(* Logix 5000 project; controller NWGG 1756-L72 rev 35.12; software revision 35.00; part 11 of 19 *)
(* tags used below, declared in another part *)
   _108M : ALIAS FOR O25[10].15;
   _109M : ALIAS FOR O25[10].9;
   _116M : ALIAS FOR O25[10].10;
   _117M : ALIAS FOR O25[10].8;
   _11_GATE_PO1 : ALIAS FOR N14[11];
   _11_GATE_PO_STOR : REAL;
   _123M : ALIAS FOR O25[10].6;
   _12_GATE_PO1 : ALIAS FOR N14[12];
   _12_GATE_PO_STOR : REAL;
   _13_GATE_PO1 : ALIAS FOR N14[13];
   _13_GATE_PO_STOR : REAL;
   _14_GATE_PO1 : ALIAS FOR N14[14];
   _14_GATE_PO_STOR : REAL;
   _15_GATE_PO1 : ALIAS FOR N14[15];
   _15_GATE_PO_STOR : REAL;
   _16_GATE_PO1 : ALIAS FOR N14[16];
   _16_GATE_PO_STOR : REAL;
   _17_GATE_PO1 : ALIAS FOR N14[17];
   _17_GATE_PO_STOR : REAL;
   _21_GATE_PO1 : ALIAS FOR N14[21];
   _21_GATE_PO_STOR : REAL;
   _22_GATE_PO1 : ALIAS FOR N14[22];
   _22_GATE_PO_STOR : REAL;
   _23_GATE_PO1 : ALIAS FOR N14[23];
   _23_GATE_PO_STOR : REAL;
   _24_GATE_PO1 : ALIAS FOR N14[24];
   _24_GATE_PO_STOR : REAL;
   _25_GATE_PO1 : ALIAS FOR N14[25];
   _25_GATE_PO_STOR : REAL;
   _26_GATE_PO1 : ALIAS FOR N14[26];
   _26_GATE_PO_STOR : REAL;
   _35M : ALIAS FOR O25[10].13;
   _43M : ALIAS FOR O25[10].14;
   _705M : ALIAS FOR O25[10].12;
   B3 : DINT[250];
   cpBinGateRates : DINT[50];
   cpBINOPEN : DINT;
   cpCleanBulk : BOOL;
   cpTicketBinActive : DINT;
   cpTicketBinSet : DINT;
   cpVAR_BINARRAY : STRING[50];
   cpVAR_CNT_ONS : DINT;
   cpVarTrimTemp : STRING;
   indexTbl : DINT;
   indexTRTTbl : DINT;
   O24 : INT[32];
   O24_007_Bit10 : ALIAS FOR O24[7].10;
   O24_007_Bit11 : ALIAS FOR O24[7].11;
   O24_007_Bit12 : ALIAS FOR O24[7].12;
   O24_007_Bit13 : ALIAS FOR O24[7].13;
   O24_007_Bit14 : ALIAS FOR O24[7].14;
   P10_RUN_AU1 : ALIAS FOR B3[4].10;
   P1_RUN_AUT1 : ALIAS FOR B3[4].1;
   P2_RUN_AUT1 : ALIAS FOR B3[4].2;
   P3_RUN_AUT1 : ALIAS FOR B3[4].3;
   P4_RUN_AUT1 : ALIAS FOR B3[4].4;
   P5_RUN_AUT1 : ALIAS FOR B3[4].5;
   P6_RUN_AUT1 : ALIAS FOR B3[4].6;
   P7_RUN_AUT1 : ALIAS FOR B3[4].7;
   P8_RUN_AUT1 : ALIAS FOR B3[4].8;
   PUMP_13_RUN : ALIAS FOR R3M1_AENTR:3:O.8;
   PUMP_14_RUN : ALIAS FOR R3M1_AENTR:3:O.9;
   PUMP_15_RUN : ALIAS FOR R3M1_AENTR:3:O.14;
   spBinGateRates : DINT[50];
   spTicketProcessing : BOOL;
   strEmptyVar : STRING;
   TicketTreatPumpActive : DINT;
   TicketTreatPumpSet : DINT;
   TRT_ARRAY : STRING[50];
   TRT_CNT : DINT;
   TRT_CNT_ONS : DINT;
   Trt_CntStore : DINT;
   TRT_PumpRATE : DINT[50];
   TRT_TICKETtable : STRING[100];
   TRT_TickettableItemNo : DINT[50];
   TRT_TICKETtableRate : DINT[100];
   TrtTrimTemp : STRING;
   VAR_CNT : DINT;
   Var_CntStore : DINT;
   VAR_TICKETtable : STRING[20];
   VAR_TickettableItemNo : DINT[50];
   VAR_TICKETtableRate : DINT[100];
   vartableONS : DINT;
   zzztmpTANKtest : DINT[10];
(* MainProgram, continued *)

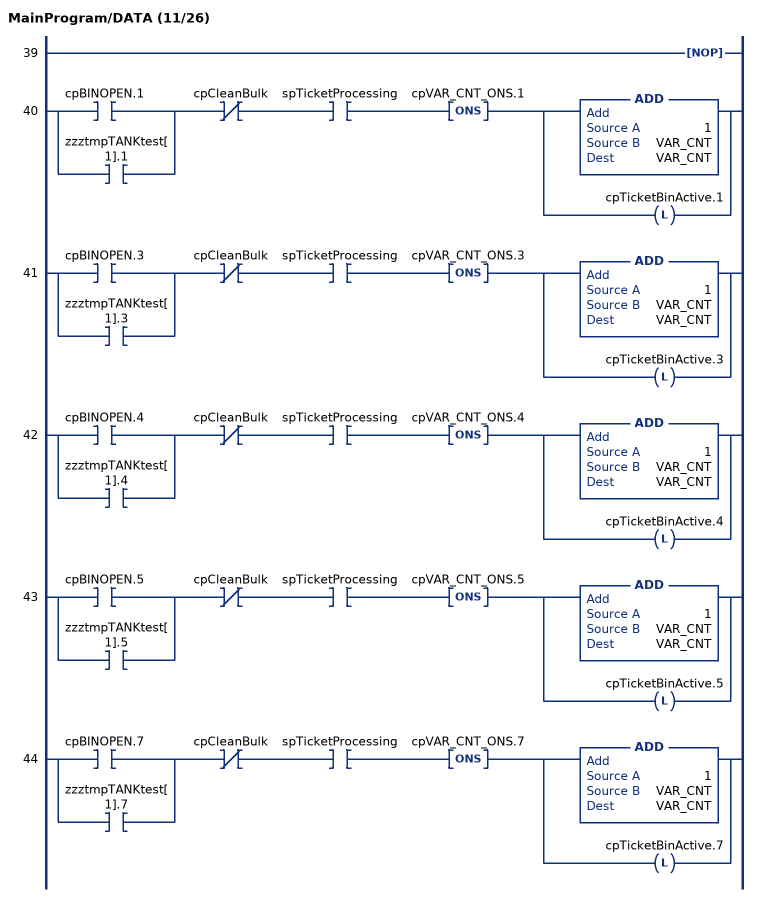
   [picture p209: MainProgram/DATA rungs 39-44]
   39: NOP();
   40: [XIC(cpBINOPEN.1) ,XIC(zzztmpTANKtest[1].1) ]XIO(cpCleanBulk)XIC(spTicketProcessing)ONS(cpVAR_CNT_ONS.1)[ADD(1,VAR_CNT,VAR_CNT) ,OTL(cpTicketBinActive.1) ];
   41: [XIC(cpBINOPEN.3) ,XIC(zzztmpTANKtest[1].3) ]XIO(cpCleanBulk)XIC(spTicketProcessing)ONS(cpVAR_CNT_ONS.3)[ADD(1,VAR_CNT,VAR_CNT) ,OTL(cpTicketBinActive.3) ];
   42: [XIC(cpBINOPEN.4) ,XIC(zzztmpTANKtest[1].4) ]XIO(cpCleanBulk)XIC(spTicketProcessing)ONS(cpVAR_CNT_ONS.4)[ADD(1,VAR_CNT,VAR_CNT) ,OTL(cpTicketBinActive.4) ];
   43: [XIC(cpBINOPEN.5) ,XIC(zzztmpTANKtest[1].5) ]XIO(cpCleanBulk)XIC(spTicketProcessing)ONS(cpVAR_CNT_ONS.5)[ADD(1,VAR_CNT,VAR_CNT) ,OTL(cpTicketBinActive.5) ];
   44: [XIC(cpBINOPEN.7) ,XIC(zzztmpTANKtest[1].7) ]XIO(cpCleanBulk)XIC(spTicketProcessing)ONS(cpVAR_CNT_ONS.7)[ADD(1,VAR_CNT,VAR_CNT) ,OTL(cpTicketBinActive.7) ];
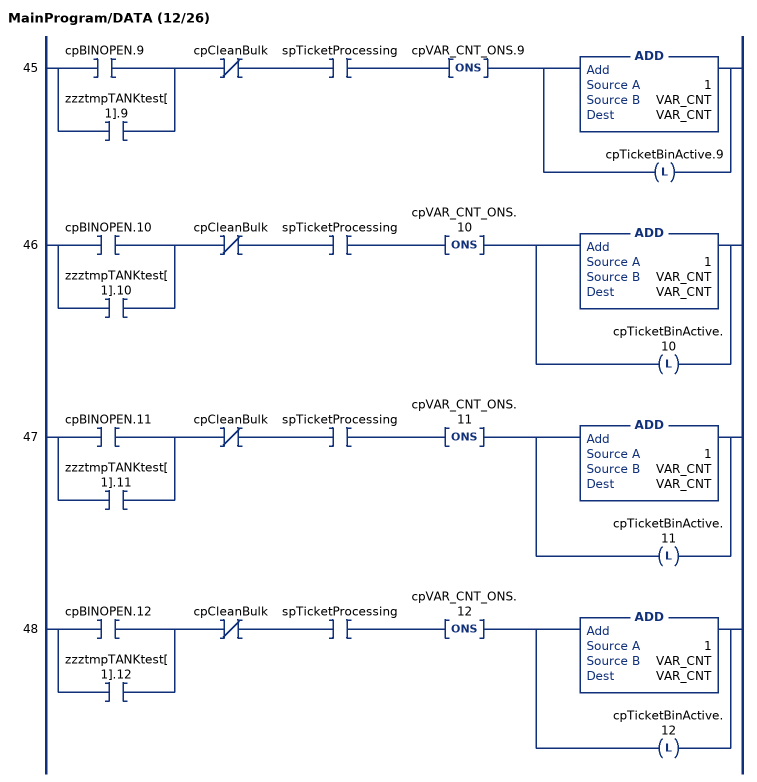
   45: [XIC(cpBINOPEN.9) ,XIC(zzztmpTANKtest[1].9) ]XIO(cpCleanBulk)XIC(spTicketProcessing)ONS(cpVAR_CNT_ONS.9)[ADD(1,VAR_CNT,VAR_CNT) ,OTL(cpTicketBinActive.9) ];
   46: [XIC(cpBINOPEN.10) ,XIC(zzztmpTANKtest[1].10) ]XIO(cpCleanBulk)XIC(spTicketProcessing)ONS(cpVAR_CNT_ONS.10)[ADD(1,VAR_CNT,VAR_CNT) ,OTL(cpTicketBinActive.10) ];
   47: [XIC(cpBINOPEN.11) ,XIC(zzztmpTANKtest[1].11) ]XIO(cpCleanBulk)XIC(spTicketProcessing)ONS(cpVAR_CNT_ONS.11)[ADD(1,VAR_CNT,VAR_CNT) ,OTL(cpTicketBinActive.11) ];
   48: [XIC(cpBINOPEN.12) ,XIC(zzztmpTANKtest[1].12) ]XIO(cpCleanBulk)XIC(spTicketProcessing)ONS(cpVAR_CNT_ONS.12)[ADD(1,VAR_CNT,VAR_CNT) ,OTL(cpTicketBinActive.12) ];
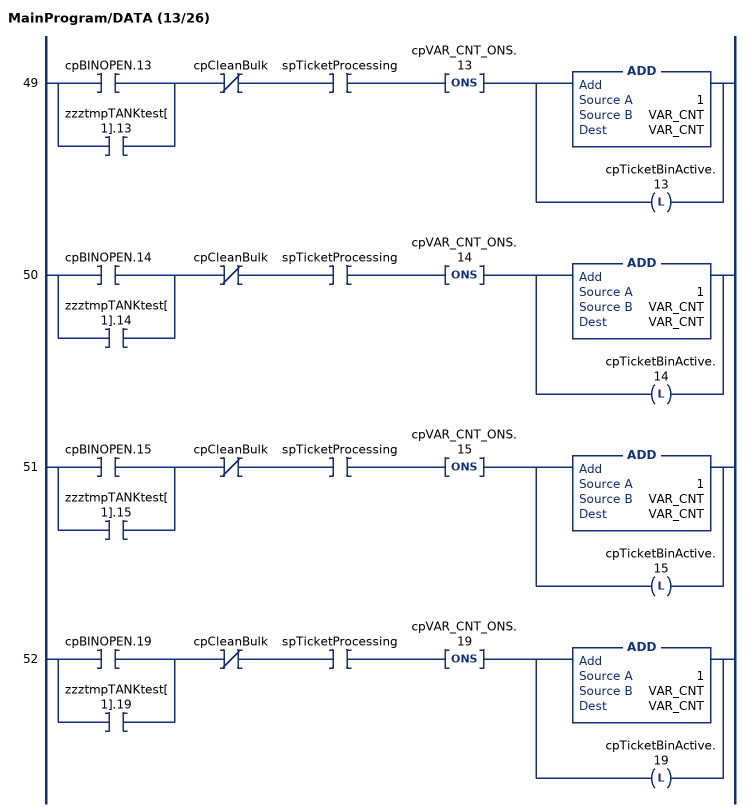
   49: [XIC(cpBINOPEN.13) ,XIC(zzztmpTANKtest[1].13) ]XIO(cpCleanBulk)XIC(spTicketProcessing)ONS(cpVAR_CNT_ONS.13)[ADD(1,VAR_CNT,VAR_CNT) ,OTL(cpTicketBinActive.13) ];
   50: [XIC(cpBINOPEN.14) ,XIC(zzztmpTANKtest[1].14) ]XIO(cpCleanBulk)XIC(spTicketProcessing)ONS(cpVAR_CNT_ONS.14)[ADD(1,VAR_CNT,VAR_CNT) ,OTL(cpTicketBinActive.14) ];
   51: [XIC(cpBINOPEN.15) ,XIC(zzztmpTANKtest[1].15) ]XIO(cpCleanBulk)XIC(spTicketProcessing)ONS(cpVAR_CNT_ONS.15)[ADD(1,VAR_CNT,VAR_CNT) ,OTL(cpTicketBinActive.15) ];
   52: [XIC(cpBINOPEN.19) ,XIC(zzztmpTANKtest[1].19) ]XIO(cpCleanBulk)XIC(spTicketProcessing)ONS(cpVAR_CNT_ONS.19)[ADD(1,VAR_CNT,VAR_CNT) ,OTL(cpTicketBinActive.19) ];
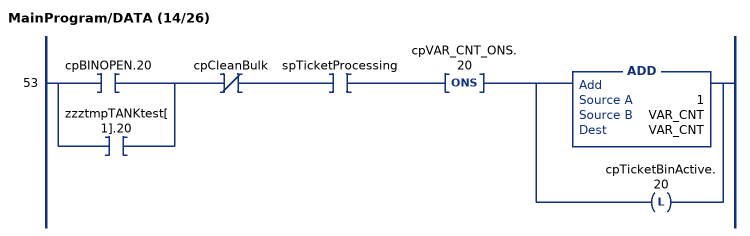
   53: [XIC(cpBINOPEN.20) ,XIC(zzztmpTANKtest[1].20) ]XIO(cpCleanBulk)XIC(spTicketProcessing)ONS(cpVAR_CNT_ONS.20)[ADD(1,VAR_CNT,VAR_CNT) ,OTL(cpTicketBinActive.20) ];
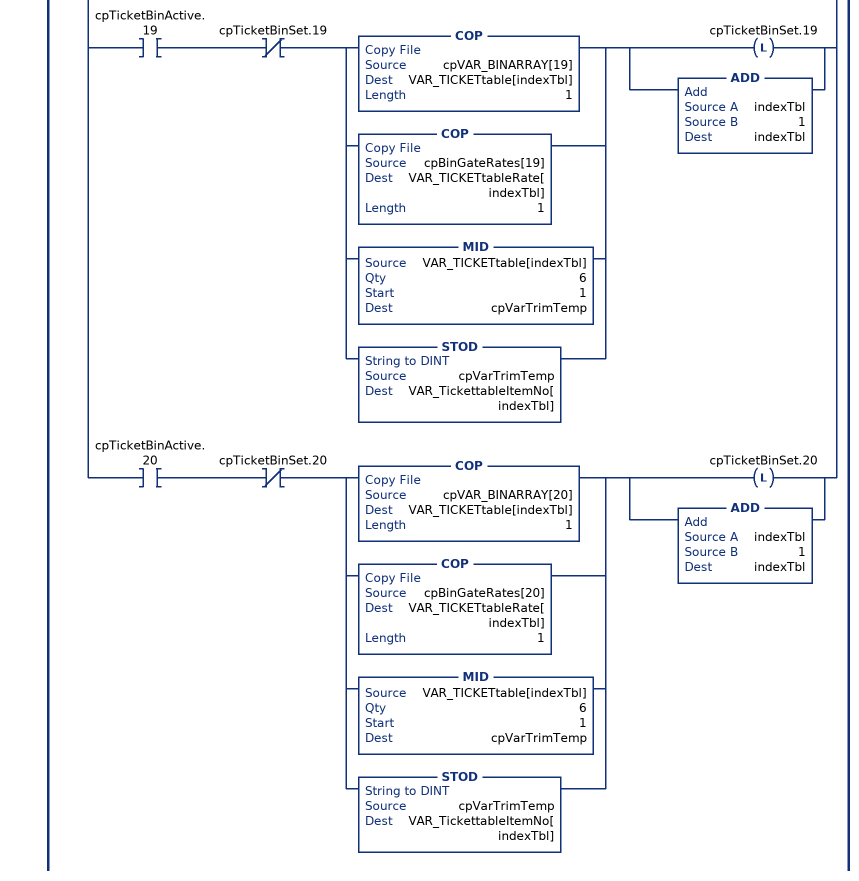
   54: GRT(VAR_CNT,0)LES(indexTbl,VAR_CNT)[XIC(cpTicketBinActive.1) XIO(cpTicketBinSet.1) [COP(cpVAR_BINARRAY[1],VAR_TICKETtable[indexTbl],1) ,COP(cpBinGateRates[1],VAR_TICKETtableRate[indexTbl],1) ,MID(VAR_TICKETtable[indexTbl],6,1,cpVarTrimTemp) ,STOD(cpVarTrimTemp,VAR_TickettableItemNo[indexTbl]) ] [OTL(cpTicketBinSet.1) ,ADD(indexTbl,1,indexTbl) ] ,XIC(cpTicketBinActive.3) XIO(cpTicketBinSet.3) [COP(cpVAR_BINARRAY[3],VAR_TICKETtable[indexTbl],1) ,COP(cpBinGateRates[3],VAR_TICKETtableRate[indexTbl],1) ,MID(VAR_TICKETtable[indexTbl],6,1,cpVarTrimTemp) ,STOD(cpVarTrimTemp,VAR_TickettableItemNo[indexTbl]) ] [OTL(cpTicketBinSet.3) ,ADD(indexTbl,1,indexTbl) ] ,XIC(cpTicketBinActive.4) XIO(cpTicketBinSet.4) [COP(cpVAR_BINARRAY[4],VAR_TICKETtable[indexTbl],1) ,COP(cpBinGateRates[4],VAR_TICKETtableRate[indexTbl],1) ,MID(VAR_TICKETtable[indexTbl],6,1,cpVarTrimTemp) ,STOD(cpVarTrimTemp,VAR_TickettableItemNo[indexTbl]) ] [OTL(cpTicketBinSet.4) ,ADD(indexTbl,1,indexTbl) ] ,XIC(cpTicketBinActive.5) XIO(cpTicketBinSet.5) [COP(cpVAR_BINARRAY[5],VAR_TICKETtable[indexTbl],1) ,COP(cpBinGateRates[5],VAR_TICKETtableRate[indexTbl],1) ,MID(VAR_TICKETtable[indexTbl],6,1,cpVarTrimTemp) ,STOD(cpVarTrimTemp,VAR_TickettableItemNo[indexTbl]) ] [OTL(cpTicketBinSet.5) ,ADD(indexTbl,1,indexTbl) ] ,XIC(cpTicketBinActive.7) XIO(cpTicketBinSet.7) [COP(cpVAR_BINARRAY[7],VAR_TICKETtable[indexTbl],1) ,COP(cpBinGateRates[7],VAR_TICKETtableRate[indexTbl],1) ,MID(VAR_TICKETtable[indexTbl],6,1,cpVarTrimTemp) ,STOD(cpVarTrimTemp,VAR_TickettableItemNo[indexTbl]) ] [OTL(cpTicketBinSet.7) ,ADD(indexTbl,1,indexTbl) ] ,XIC(cpTicketBinActive.9) XIO(cpTicketBinSet.9) [COP(cpVAR_BINARRAY[9],VAR_TICKETtable[indexTbl],1) ,COP(cpBinGateRates[9],VAR_TICKETtableRate[indexTbl],1) ,MID(VAR_TICKETtable[indexTbl],6,1,cpVarTrimTemp) ,STOD(cpVarTrimTemp,VAR_TickettableItemNo[indexTbl]) ] [OTL(cpTicketBinSet.9) ,ADD(indexTbl,1,indexTbl) ] ,XIC(cpTicketBinActive.10) XIO(cpTicketBinSet.10) [COP(cpVAR_BINARRAY[10],VAR_TICKETtable[indexTbl],1) ,COP(cpBinGateRates[10],VAR_TICKETtableRate[indexTbl],1) ,MID(VAR_TICKETtable[indexTbl],6,1,cpVarTrimTemp) ,STOD(cpVarTrimTemp,VAR_TickettableItemNo[indexTbl]) ] [OTL(cpTicketBinSet.10) ,ADD(indexTbl,1,indexTbl) ] ,XIC(cpTicketBinActive.11) XIO(cpTicketBinSet.11) [COP(cpVAR_BINARRAY[11],VAR_TICKETtable[indexTbl],1) ,COP(cpBinGateRates[11],VAR_TICKETtableRate[indexTbl],1) ,MID(VAR_TICKETtable[indexTbl],6,1,cpVarTrimTemp) ,STOD(cpVarTrimTemp,VAR_TickettableItemNo[indexTbl]) ] [OTL(cpTicketBinSet.11) ,ADD(indexTbl,1,indexTbl) ] ,XIC(cpTicketBinActive.12) XIO(cpTicketBinSet.12) [COP(cpVAR_BINARRAY[12],VAR_TICKETtable[indexTbl],1) ,COP(cpBinGateRates[12],VAR_TICKETtableRate[indexTbl],1) ,MID(VAR_TICKETtable[indexTbl],6,1,cpVarTrimTemp) ,STOD(cpVarTrimTemp,VAR_TickettableItemNo[indexTbl]) ] [OTL(cpTicketBinSet.12) ,ADD(indexTbl,1,indexTbl) ] ,XIC(cpTicketBinActive.13) XIO(cpTicketBinSet.13) [COP(cpVAR_BINARRAY[13],VAR_TICKETtable[indexTbl],1) ,COP(cpBinGateRates[13],VAR_TICKETtableRate[indexTbl],1) ,MID(VAR_TICKETtable[indexTbl],6,1,cpVarTrimTemp) ,STOD(cpVarTrimTemp,VAR_TickettableItemNo[indexTbl]) ] [OTL(cpTicketBinSet.13) ,ADD(indexTbl,1,indexTbl) ] ,XIC(cpTicketBinActive.14) XIO(cpTicketBinSet.14) [COP(cpVAR_BINARRAY[14],VAR_TICKETtable[indexTbl],1) ,COP(cpBinGateRates[14],VAR_TICKETtableRate[indexTbl],1) ,MID(VAR_TICKETtable[indexTbl],6,1,cpVarTrimTemp) ,STOD(cpVarTrimTemp,VAR_TickettableItemNo[indexTbl]) ] [OTL(cpTicketBinSet.14) ,ADD(indexTbl,1,indexTbl) ] ,XIC(cpTicketBinActive.15) XIO(cpTicketBinSet.15) [COP(cpVAR_BINARRAY[15],VAR_TICKETtable[indexTbl],1) ,COP(cpBinGateRates[15],VAR_TICKETtableRate[indexTbl],1) ,MID(VAR_TICKETtable[indexTbl],6,1,cpVarTrimTemp) ,STOD(cpVarTrimTemp,VAR_TickettableItemNo[indexTbl]) ] [OTL(cpTicketBinSet.15) ,ADD(indexTbl,1,indexTbl) ] ,XIC(cpTicketBinActive.19) XIO(cpTicketBinSet.19) [COP(cpVAR_BINARRAY[19],VAR_TICKETtable[indexTbl],1) ,COP(cpBinGateRates[19],VAR_TICKETtableRate[indexTbl],1) ,MID(VAR_TICKETtable[indexTbl],6,1,cpVarTrimTemp) ,STOD(cpVarTrimTemp,VAR_TickettableItemNo[indexTbl]) ] [OTL(cpTicketBinSet.19) ,ADD(indexTbl,1,indexTbl) ] ,XIC(cpTicketBinActive.20) XIO(cpTicketBinSet.20) [COP(cpVAR_BINARRAY[20],VAR_TICKETtable[indexTbl],1) ,COP(cpBinGateRates[20],VAR_TICKETtableRate[indexTbl],1) ,MID(VAR_TICKETtable[indexTbl],6,1,cpVarTrimTemp) ,STOD(cpVarTrimTemp,VAR_TickettableItemNo[indexTbl]) ] [OTL(cpTicketBinSet.20) ,ADD(indexTbl,1,indexTbl) ] ];
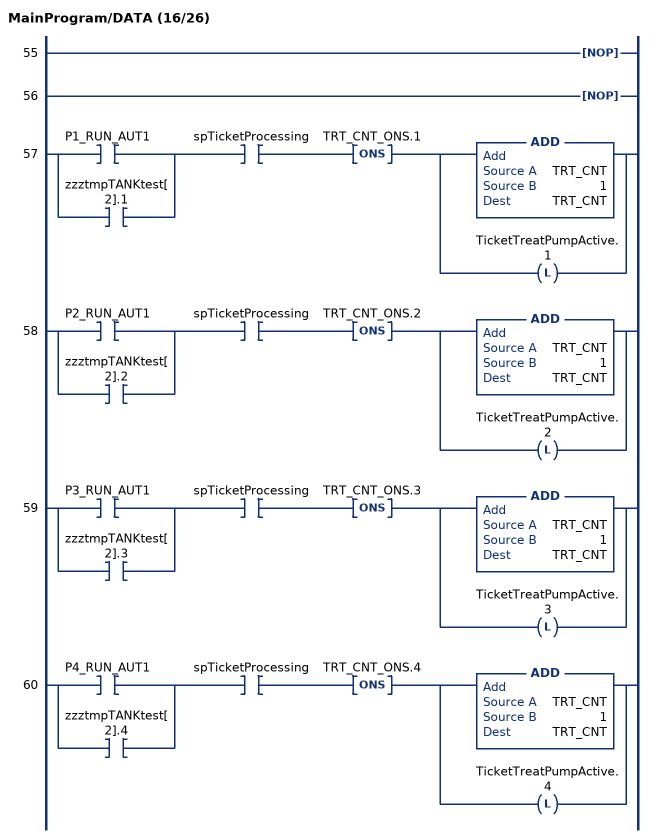
   55: NOP();
   56: NOP();
   57: [XIC(P1_RUN_AUT1) ,XIC(zzztmpTANKtest[2].1) ]XIC(spTicketProcessing)ONS(TRT_CNT_ONS.1)[ADD(TRT_CNT,1,TRT_CNT) ,OTL(TicketTreatPumpActive.1) ];
   58: [XIC(P2_RUN_AUT1) ,XIC(zzztmpTANKtest[2].2) ]XIC(spTicketProcessing)ONS(TRT_CNT_ONS.2)[ADD(TRT_CNT,1,TRT_CNT) ,OTL(TicketTreatPumpActive.2) ];
   59: [XIC(P3_RUN_AUT1) ,XIC(zzztmpTANKtest[2].3) ]XIC(spTicketProcessing)ONS(TRT_CNT_ONS.3)[ADD(TRT_CNT,1,TRT_CNT) ,OTL(TicketTreatPumpActive.3) ];
   60: [XIC(P4_RUN_AUT1) ,XIC(zzztmpTANKtest[2].4) ]XIC(spTicketProcessing)ONS(TRT_CNT_ONS.4)[ADD(TRT_CNT,1,TRT_CNT) ,OTL(TicketTreatPumpActive.4) ];
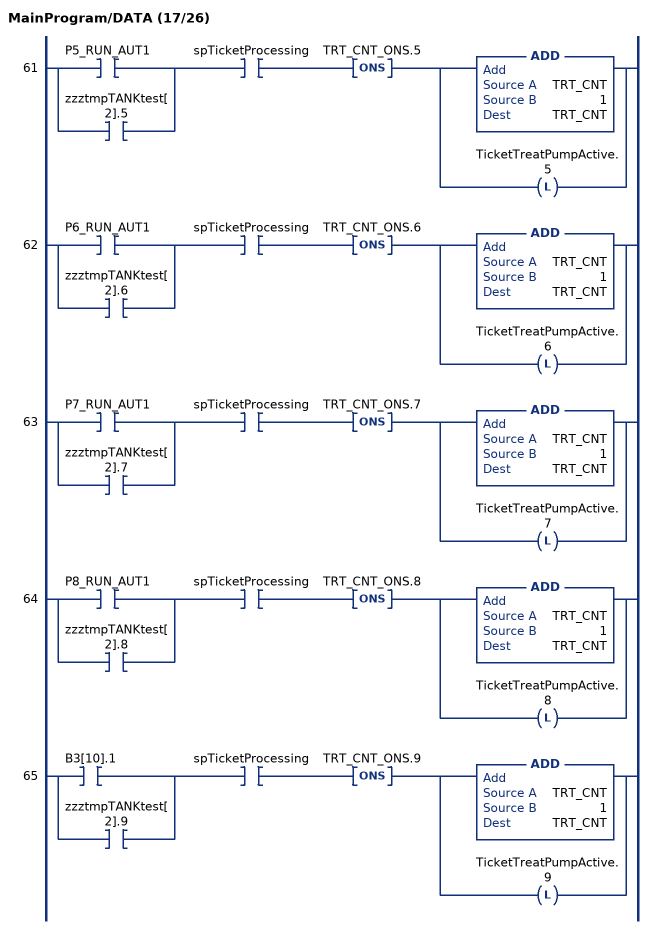
   61: [XIC(P5_RUN_AUT1) ,XIC(zzztmpTANKtest[2].5) ]XIC(spTicketProcessing)ONS(TRT_CNT_ONS.5)[ADD(TRT_CNT,1,TRT_CNT) ,OTL(TicketTreatPumpActive.5) ];
   62: [XIC(P6_RUN_AUT1) ,XIC(zzztmpTANKtest[2].6) ]XIC(spTicketProcessing)ONS(TRT_CNT_ONS.6)[ADD(TRT_CNT,1,TRT_CNT) ,OTL(TicketTreatPumpActive.6) ];
   63: [XIC(P7_RUN_AUT1) ,XIC(zzztmpTANKtest[2].7) ]XIC(spTicketProcessing)ONS(TRT_CNT_ONS.7)[ADD(TRT_CNT,1,TRT_CNT) ,OTL(TicketTreatPumpActive.7) ];
   64: [XIC(P8_RUN_AUT1) ,XIC(zzztmpTANKtest[2].8) ]XIC(spTicketProcessing)ONS(TRT_CNT_ONS.8)[ADD(TRT_CNT,1,TRT_CNT) ,OTL(TicketTreatPumpActive.8) ];
   65: [XIC(B3[10].1) ,XIC(zzztmpTANKtest[2].9) ]XIC(spTicketProcessing)ONS(TRT_CNT_ONS.9)[ADD(TRT_CNT,1,TRT_CNT) ,OTL(TicketTreatPumpActive.9) ];
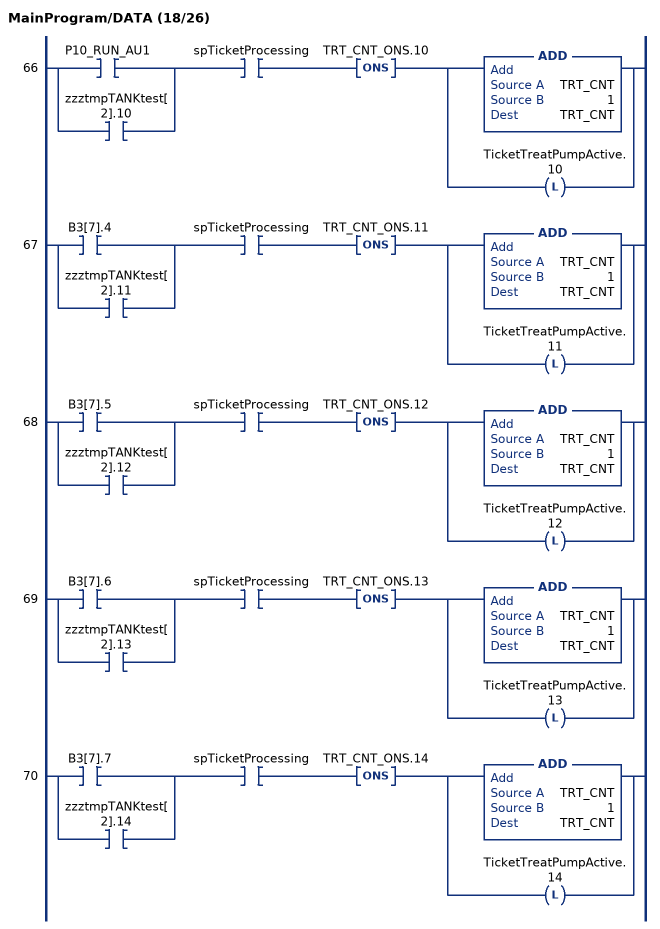
   66: [XIC(P10_RUN_AU1) ,XIC(zzztmpTANKtest[2].10) ]XIC(spTicketProcessing)ONS(TRT_CNT_ONS.10)[ADD(TRT_CNT,1,TRT_CNT) ,OTL(TicketTreatPumpActive.10) ];
   67: [XIC(B3[7].4) ,XIC(zzztmpTANKtest[2].11) ]XIC(spTicketProcessing)ONS(TRT_CNT_ONS.11)[ADD(TRT_CNT,1,TRT_CNT) ,OTL(TicketTreatPumpActive.11) ];
   68: [XIC(B3[7].5) ,XIC(zzztmpTANKtest[2].12) ]XIC(spTicketProcessing)ONS(TRT_CNT_ONS.12)[ADD(TRT_CNT,1,TRT_CNT) ,OTL(TicketTreatPumpActive.12) ];
   69: [XIC(B3[7].6) ,XIC(zzztmpTANKtest[2].13) ]XIC(spTicketProcessing)ONS(TRT_CNT_ONS.13)[ADD(TRT_CNT,1,TRT_CNT) ,OTL(TicketTreatPumpActive.13) ];
   70: [XIC(B3[7].7) ,XIC(zzztmpTANKtest[2].14) ]XIC(spTicketProcessing)ONS(TRT_CNT_ONS.14)[ADD(TRT_CNT,1,TRT_CNT) ,OTL(TicketTreatPumpActive.14) ];
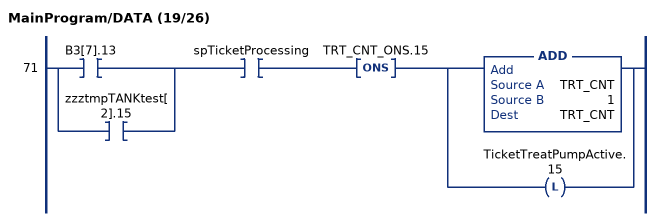
   71: [XIC(B3[7].13) ,XIC(zzztmpTANKtest[2].15) ]XIC(spTicketProcessing)ONS(TRT_CNT_ONS.15)[ADD(TRT_CNT,1,TRT_CNT) ,OTL(TicketTreatPumpActive.15) ];
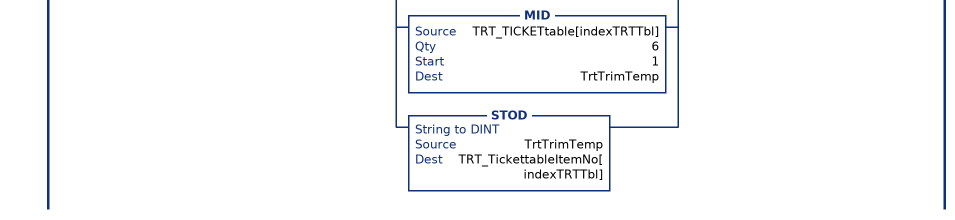
   72: GRT(TRT_CNT,0)LES(indexTRTTbl,TRT_CNT)[XIC(TicketTreatPumpActive.1) XIO(TicketTreatPumpSet.1) [COP(TRT_ARRAY[1],TRT_TICKETtable[indexTRTTbl],1) ,COP(TRT_PumpRATE[1],TRT_TICKETtableRate[indexTRTTbl],1) ,MID(TRT_TICKETtable[indexTRTTbl],6,1,TrtTrimTemp) ,STOD(TrtTrimTemp,TRT_TickettableItemNo[indexTRTTbl]) ] [OTL(TicketTreatPumpSet.1) ,ADD(indexTRTTbl,1,indexTRTTbl) ] ,XIC(TicketTreatPumpActive.2) XIO(TicketTreatPumpSet.2) [COP(TRT_ARRAY[2],TRT_TICKETtable[indexTRTTbl],1) ,COP(TRT_PumpRATE[2],TRT_TICKETtableRate[indexTRTTbl],1) ,MID(TRT_TICKETtable[indexTRTTbl],6,1,TrtTrimTemp) ,STOD(TrtTrimTemp,TRT_TickettableItemNo[indexTRTTbl]) ] [OTL(TicketTreatPumpSet.2) ,ADD(indexTRTTbl,1,indexTRTTbl) ] ,XIC(TicketTreatPumpActive.3) XIO(TicketTreatPumpSet.3) [COP(TRT_ARRAY[3],TRT_TICKETtable[indexTRTTbl],1) ,COP(TRT_PumpRATE[3],TRT_TICKETtableRate[indexTRTTbl],1) ,MID(TRT_TICKETtable[indexTRTTbl],6,1,TrtTrimTemp) ,STOD(TrtTrimTemp,TRT_TickettableItemNo[indexTRTTbl]) ] [OTL(TicketTreatPumpSet.3) ,ADD(indexTRTTbl,1,indexTRTTbl) ] ,XIC(TicketTreatPumpActive.4) XIO(TicketTreatPumpSet.4) [COP(TRT_ARRAY[4],TRT_TICKETtable[indexTRTTbl],1) ,COP(TRT_PumpRATE[4],TRT_TICKETtableRate[indexTRTTbl],1) ,MID(TRT_TICKETtable[indexTRTTbl],6,1,TrtTrimTemp) ,STOD(TrtTrimTemp,TRT_TickettableItemNo[indexTRTTbl]) ] [OTL(TicketTreatPumpSet.4) ,ADD(indexTRTTbl,1,indexTRTTbl) ] ,XIC(TicketTreatPumpActive.5) XIO(TicketTreatPumpSet.5) [COP(TRT_ARRAY[5],TRT_TICKETtable[indexTRTTbl],1) ,COP(TRT_PumpRATE[5],TRT_TICKETtableRate[indexTRTTbl],1) ,MID(TRT_TICKETtable[indexTRTTbl],6,1,TrtTrimTemp) ,STOD(TrtTrimTemp,TRT_TickettableItemNo[indexTRTTbl]) ] [OTL(TicketTreatPumpSet.5) ,ADD(indexTRTTbl,1,indexTRTTbl) ] ,XIC(TicketTreatPumpActive.6) XIO(TicketTreatPumpSet.6) [COP(TRT_ARRAY[6],TRT_TICKETtable[indexTRTTbl],1) ,COP(TRT_PumpRATE[6],TRT_TICKETtableRate[indexTRTTbl],1) ,MID(TRT_TICKETtable[indexTRTTbl],6,1,TrtTrimTemp) ,STOD(TrtTrimTemp,TRT_TickettableItemNo[indexTRTTbl]) ] [OTL(TicketTreatPumpSet.6) ,ADD(indexTRTTbl,1,indexTRTTbl) ] ,XIC(TicketTreatPumpActive.7) XIO(TicketTreatPumpSet.7) [COP(TRT_ARRAY[7],TRT_TICKETtable[indexTRTTbl],1) ,COP(TRT_PumpRATE[7],TRT_TICKETtableRate[indexTRTTbl],1) ,MID(TRT_TICKETtable[indexTRTTbl],6,1,TrtTrimTemp) ,STOD(TrtTrimTemp,TRT_TickettableItemNo[indexTRTTbl]) ] [OTL(TicketTreatPumpSet.7) ,ADD(indexTRTTbl,1,indexTRTTbl) ] ,XIC(TicketTreatPumpActive.8) XIO(TicketTreatPumpSet.8) [COP(TRT_ARRAY[8],TRT_TICKETtable[indexTRTTbl],1) ,COP(TRT_PumpRATE[8],TRT_TICKETtableRate[indexTRTTbl],1) ,MID(TRT_TICKETtable[indexTRTTbl],6,1,TrtTrimTemp) ,STOD(TrtTrimTemp,TRT_TickettableItemNo[indexTRTTbl]) ] [OTL(TicketTreatPumpSet.8) ,ADD(indexTRTTbl,1,indexTRTTbl) ] ,XIC(TicketTreatPumpActive.9) XIO(TicketTreatPumpSet.9) [COP(TRT_ARRAY[9],TRT_TICKETtable[indexTRTTbl],1) ,COP(TRT_PumpRATE[9],TRT_TICKETtableRate[indexTRTTbl],1) ,MID(TRT_TICKETtable[indexTRTTbl],6,1,TrtTrimTemp) ,STOD(TrtTrimTemp,TRT_TickettableItemNo[indexTRTTbl]) ] [OTL(TicketTreatPumpSet.9) ,ADD(indexTRTTbl,1,indexTRTTbl) ] ,XIC(TicketTreatPumpActive.10) XIO(TicketTreatPumpSet.10) [COP(TRT_ARRAY[10],TRT_TICKETtable[indexTRTTbl],1) ,COP(TRT_PumpRATE[10],TRT_TICKETtableRate[indexTRTTbl],1) ,MID(TRT_TICKETtable[indexTRTTbl],6,1,TrtTrimTemp) ,STOD(TrtTrimTemp,TRT_TickettableItemNo[indexTRTTbl]) ] [OTL(TicketTreatPumpSet.10) ,ADD(indexTRTTbl,1,indexTRTTbl) ] ,XIC(TicketTreatPumpActive.11) XIO(TicketTreatPumpSet.11) [COP(TRT_ARRAY[11],TRT_TICKETtable[indexTRTTbl],1) ,COP(TRT_PumpRATE[11],TRT_TICKETtableRate[indexTRTTbl],1) ,MID(TRT_TICKETtable[indexTRTTbl],6,1,TrtTrimTemp) ,STOD(TrtTrimTemp,TRT_TickettableItemNo[indexTRTTbl]) ] [OTL(TicketTreatPumpSet.11) ,ADD(indexTRTTbl,1,indexTRTTbl) ] ,XIC(TicketTreatPumpActive.12) XIO(TicketTreatPumpSet.12) [COP(TRT_ARRAY[12],TRT_TICKETtable[indexTRTTbl],1) ,COP(TRT_PumpRATE[12],TRT_TICKETtableRate[indexTRTTbl],1) ,MID(TRT_TICKETtable[indexTRTTbl],6,1,TrtTrimTemp) ,STOD(TrtTrimTemp,TRT_TickettableItemNo[indexTRTTbl]) ] [OTL(TicketTreatPumpSet.12) ,ADD(indexTRTTbl,1,indexTRTTbl) ] ,XIC(TicketTreatPumpActive.13) XIO(TicketTreatPumpSet.13) [COP(TRT_ARRAY[13],TRT_TICKETtable[indexTRTTbl],1) ,COP(TRT_PumpRATE[14],TRT_TICKETtableRate[indexTRTTbl],1) ,MID(TRT_TICKETtable[indexTRTTbl],6,1,TrtTrimTemp) ,STOD(TrtTrimTemp,TRT_TickettableItemNo[indexTRTTbl]) ] [OTL(TicketTreatPumpSet.13) ,ADD(indexTRTTbl,1,indexTRTTbl) ] ,XIC(TicketTreatPumpActive.14) XIO(TicketTreatPumpSet.14) [COP(TRT_ARRAY[14],TRT_TICKETtable[indexTRTTbl],1) ,COP(TRT_PumpRATE[14],TRT_TICKETtableRate[indexTRTTbl],1) ,MID(TRT_TICKETtable[indexTRTTbl],6,1,TrtTrimTemp) ,STOD(TrtTrimTemp,TRT_TickettableItemNo[indexTRTTbl]) ] [OTL(TicketTreatPumpSet.14) ,ADD(indexTRTTbl,1,indexTRTTbl) ] ,XIC(TicketTreatPumpActive.15) XIO(TicketTreatPumpSet.15) [COP(TRT_ARRAY[15],TRT_TICKETtable[indexTRTTbl],1) ,COP(TRT_PumpRATE[15],TRT_TICKETtableRate[indexTRTTbl],1) ,MID(TRT_TICKETtable[indexTRTTbl],6,1,TrtTrimTemp) ,STOD(TrtTrimTemp,TRT_TickettableItemNo[indexTRTTbl]) ] [OTL(TicketTreatPumpSet.15) ,ADD(indexTRTTbl,1,indexTRTTbl) ] ];
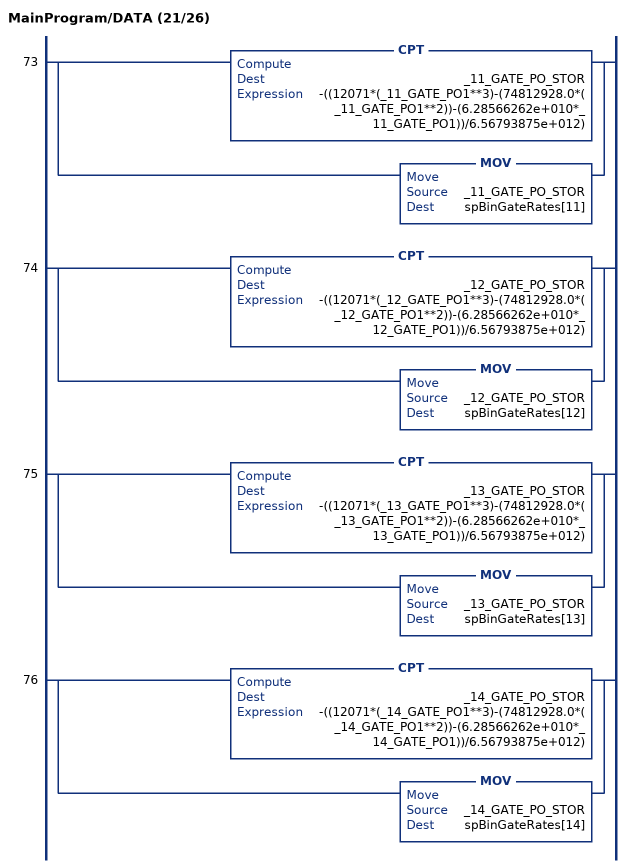
   73: [CPT(_11_GATE_PO_STOR,-((12071*(_11_GATE_PO1**3)-(74812928.0*(_11_GATE_PO1**2))-(6.28566262e+010*_11_GATE_PO1))/6.56793875e+012)) ,MOV(_11_GATE_PO_STOR,spBinGateRates[11]) ];
   74: [CPT(_12_GATE_PO_STOR,-((12071*(_12_GATE_PO1**3)-(74812928.0*(_12_GATE_PO1**2))-(6.28566262e+010*_12_GATE_PO1))/6.56793875e+012)) ,MOV(_12_GATE_PO_STOR,spBinGateRates[12]) ];
   75: [CPT(_13_GATE_PO_STOR,-((12071*(_13_GATE_PO1**3)-(74812928.0*(_13_GATE_PO1**2))-(6.28566262e+010*_13_GATE_PO1))/6.56793875e+012)) ,MOV(_13_GATE_PO_STOR,spBinGateRates[13]) ];
   76: [CPT(_14_GATE_PO_STOR,-((12071*(_14_GATE_PO1**3)-(74812928.0*(_14_GATE_PO1**2))-(6.28566262e+010*_14_GATE_PO1))/6.56793875e+012)) ,MOV(_14_GATE_PO_STOR,spBinGateRates[14]) ];
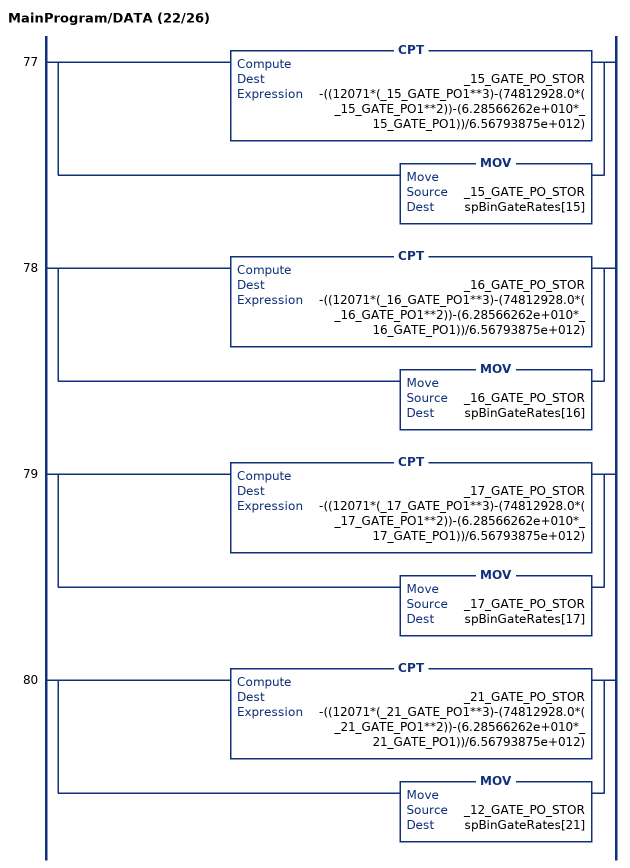
   77: [CPT(_15_GATE_PO_STOR,-((12071*(_15_GATE_PO1**3)-(74812928.0*(_15_GATE_PO1**2))-(6.28566262e+010*_15_GATE_PO1))/6.56793875e+012)) ,MOV(_15_GATE_PO_STOR,spBinGateRates[15]) ];
   78: [CPT(_16_GATE_PO_STOR,-((12071*(_16_GATE_PO1**3)-(74812928.0*(_16_GATE_PO1**2))-(6.28566262e+010*_16_GATE_PO1))/6.56793875e+012)) ,MOV(_16_GATE_PO_STOR,spBinGateRates[16]) ];
   79: [CPT(_17_GATE_PO_STOR,-((12071*(_17_GATE_PO1**3)-(74812928.0*(_17_GATE_PO1**2))-(6.28566262e+010*_17_GATE_PO1))/6.56793875e+012)) ,MOV(_17_GATE_PO_STOR,spBinGateRates[17]) ];
   80: [CPT(_21_GATE_PO_STOR,-((12071*(_21_GATE_PO1**3)-(74812928.0*(_21_GATE_PO1**2))-(6.28566262e+010*_21_GATE_PO1))/6.56793875e+012)) ,MOV(_12_GATE_PO_STOR,spBinGateRates[21]) ];
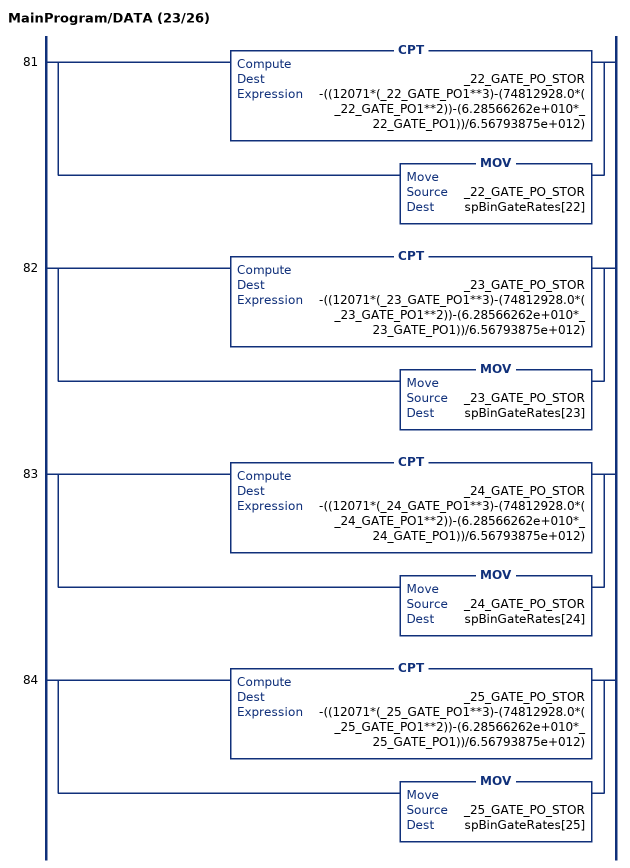
   81: [CPT(_22_GATE_PO_STOR,-((12071*(_22_GATE_PO1**3)-(74812928.0*(_22_GATE_PO1**2))-(6.28566262e+010*_22_GATE_PO1))/6.56793875e+012)) ,MOV(_22_GATE_PO_STOR,spBinGateRates[22]) ];
   82: [CPT(_23_GATE_PO_STOR,-((12071*(_23_GATE_PO1**3)-(74812928.0*(_23_GATE_PO1**2))-(6.28566262e+010*_23_GATE_PO1))/6.56793875e+012)) ,MOV(_23_GATE_PO_STOR,spBinGateRates[23]) ];
   83: [CPT(_24_GATE_PO_STOR,-((12071*(_24_GATE_PO1**3)-(74812928.0*(_24_GATE_PO1**2))-(6.28566262e+010*_24_GATE_PO1))/6.56793875e+012)) ,MOV(_24_GATE_PO_STOR,spBinGateRates[24]) ];
   84: [CPT(_25_GATE_PO_STOR,-((12071*(_25_GATE_PO1**3)-(74812928.0*(_25_GATE_PO1**2))-(6.28566262e+010*_25_GATE_PO1))/6.56793875e+012)) ,MOV(_25_GATE_PO_STOR,spBinGateRates[25]) ];
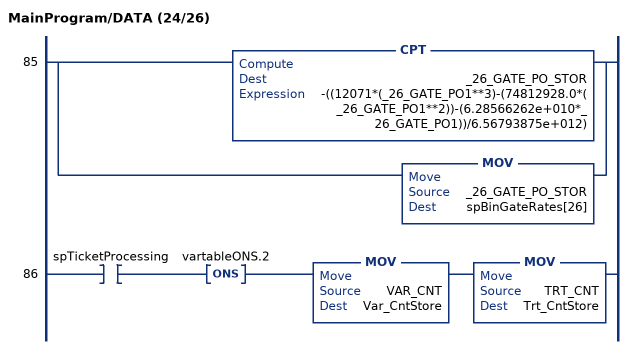
   85: [CPT(_26_GATE_PO_STOR,-((12071*(_26_GATE_PO1**3)-(74812928.0*(_26_GATE_PO1**2))-(6.28566262e+010*_26_GATE_PO1))/6.56793875e+012)) ,MOV(_26_GATE_PO_STOR,spBinGateRates[26]) ];
   86: XIC(spTicketProcessing)ONS(vartableONS.2)MOV(VAR_CNT,Var_CntStore)MOV(TRT_CNT,Trt_CntStore);
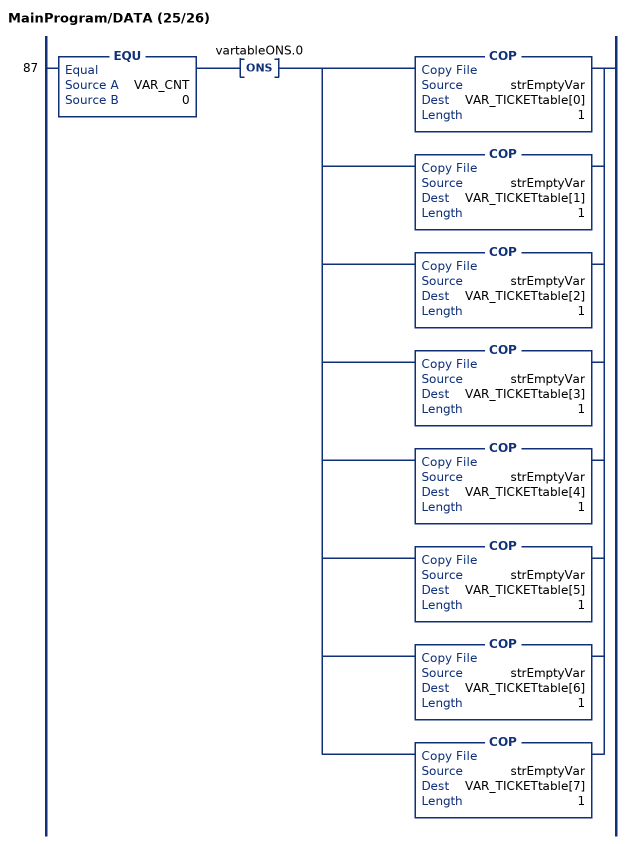
   87: EQU(VAR_CNT,0)ONS(vartableONS.0)[COP(strEmptyVar,VAR_TICKETtable[0],1) ,COP(strEmptyVar,VAR_TICKETtable[1],1) ,COP(strEmptyVar,VAR_TICKETtable[2],1) ,COP(strEmptyVar,VAR_TICKETtable[3],1) ,COP(strEmptyVar,VAR_TICKETtable[4],1) ,COP(strEmptyVar,VAR_TICKETtable[5],1) ,COP(strEmptyVar,VAR_TICKETtable[6],1) ,COP(strEmptyVar,VAR_TICKETtable[7],1) ];
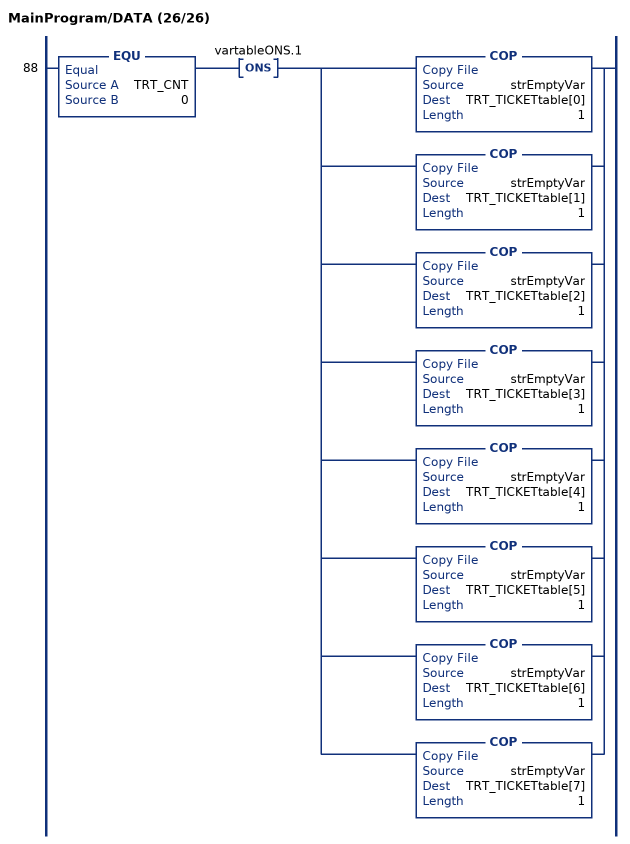
   88: EQU(TRT_CNT,0)ONS(vartableONS.1)[COP(strEmptyVar,TRT_TICKETtable[0],1) ,COP(strEmptyVar,TRT_TICKETtable[1],1) ,COP(strEmptyVar,TRT_TICKETtable[2],1) ,COP(strEmptyVar,TRT_TICKETtable[3],1) ,COP(strEmptyVar,TRT_TICKETtable[4],1) ,COP(strEmptyVar,TRT_TICKETtable[5],1) ,COP(strEmptyVar,TRT_TICKETtable[6],1) ,COP(strEmptyVar,TRT_TICKETtable[7],1) ];
END_ROUTINE

ROUTINE Dev_O24_7   (* ladder *)
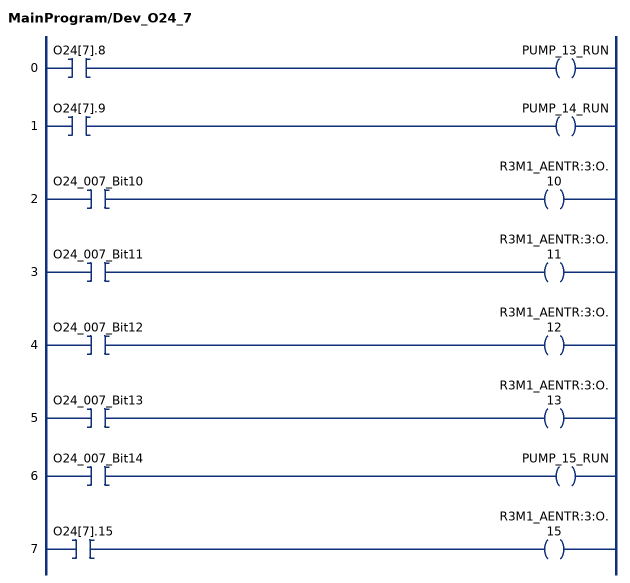
   0: XIC(O24[7].8)OTE(PUMP_13_RUN);
   1: XIC(O24[7].9)OTE(PUMP_14_RUN);
   2: XIC(O24_007_Bit10)OTE(R3M1_AENTR:3:O.10);
   3: XIC(O24_007_Bit11)OTE(R3M1_AENTR:3:O.11);
   4: XIC(O24_007_Bit12)OTE(R3M1_AENTR:3:O.12);
   5: XIC(O24_007_Bit13)OTE(R3M1_AENTR:3:O.13);
   6: XIC(O24_007_Bit14)OTE(PUMP_15_RUN);
   7: XIC(O24[7].15)OTE(R3M1_AENTR:3:O.15);
END_ROUTINE

ROUTINE Dev_O25_10   (* ladder *)
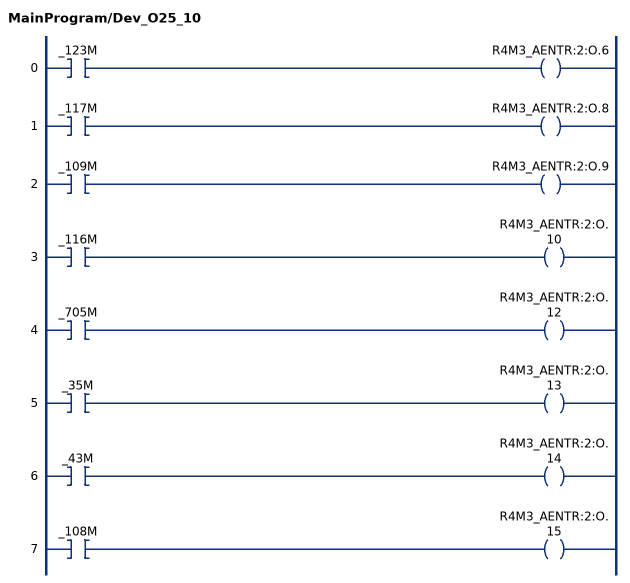
   0: XIC(_123M)OTE(R4M3_AENTR:2:O.6);
   1: XIC(_117M)OTE(R4M3_AENTR:2:O.8);
   2: XIC(_109M)OTE(R4M3_AENTR:2:O.9);
   3: XIC(_116M)OTE(R4M3_AENTR:2:O.10);
   4: XIC(_705M)OTE(R4M3_AENTR:2:O.12);
   5: XIC(_35M)OTE(R4M3_AENTR:2:O.13);
   6: XIC(_43M)OTE(R4M3_AENTR:2:O.14);
   7: XIC(_108M)OTE(R4M3_AENTR:2:O.15);
END_ROUTINE
